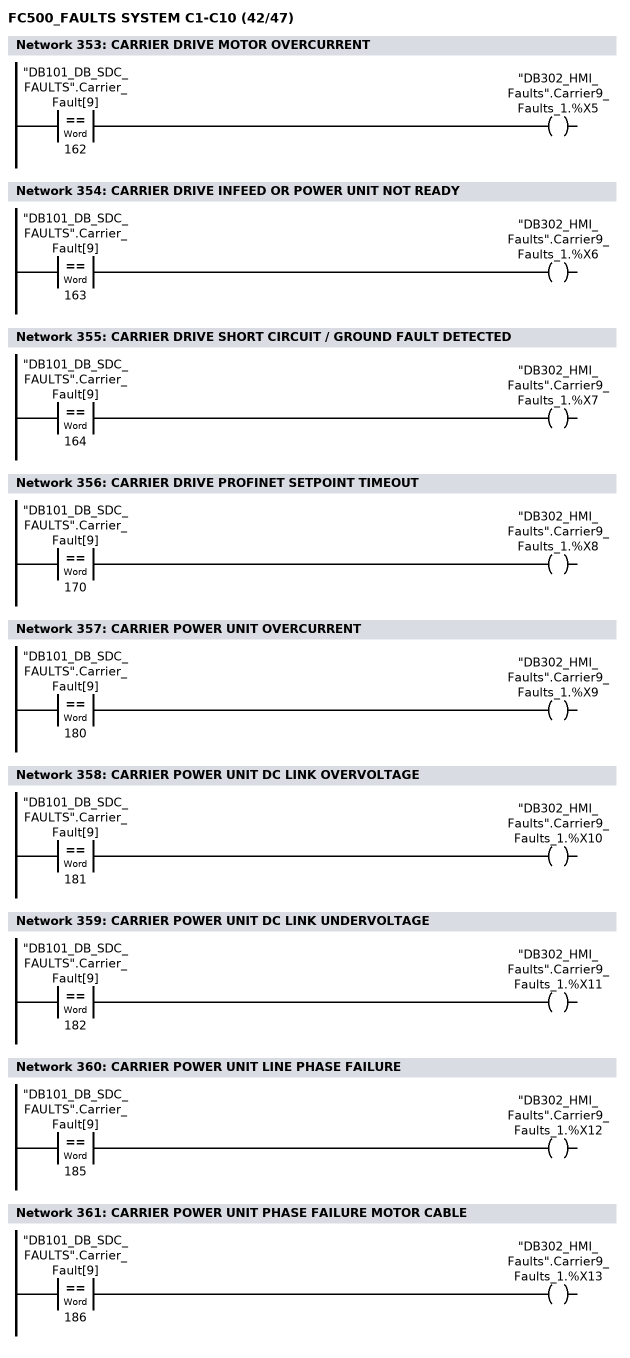
   RUNG wire#powerrail
      { S7_Templates := "SrcType := Word" } EQ_Contact(in1 := "DB101_DB_SDC_FAULTS".Carrier_Fault[9], in2 := 162)
      Coil( "DB302_HMI_Faults".Carrier9_Faults_1.%X5 )
   END_RUNG
   // the same network as SCL:
   "DB302_HMI_Faults".Carrier9_Faults_1.%X5 := "DB101_DB_SDC_FAULTS".Carrier_Fault[9] = 162;
END_REGION

REGION Network 354: CARRIER DRIVE INFEED OR POWER UNIT NOT READY
   RUNG wire#powerrail
      { S7_Templates := "SrcType := Word" } EQ_Contact(in1 := "DB101_DB_SDC_FAULTS".Carrier_Fault[9], in2 := 163)
      Coil( "DB302_HMI_Faults".Carrier9_Faults_1.%X6 )
   END_RUNG
   // the same network as SCL:
   "DB302_HMI_Faults".Carrier9_Faults_1.%X6 := "DB101_DB_SDC_FAULTS".Carrier_Fault[9] = 163;
END_REGION

REGION Network 355: CARRIER DRIVE SHORT CIRCUIT / GROUND FAULT DETECTED
   RUNG wire#powerrail
      { S7_Templates := "SrcType := Word" } EQ_Contact(in1 := "DB101_DB_SDC_FAULTS".Carrier_Fault[9], in2 := 164)
      Coil( "DB302_HMI_Faults".Carrier9_Faults_1.%X7 )
   END_RUNG
   // the same network as SCL:
   "DB302_HMI_Faults".Carrier9_Faults_1.%X7 := "DB101_DB_SDC_FAULTS".Carrier_Fault[9] = 164;
END_REGION

REGION Network 356: CARRIER DRIVE PROFINET SETPOINT TIMEOUT
   RUNG wire#powerrail
      { S7_Templates := "SrcType := Word" } EQ_Contact(in1 := "DB101_DB_SDC_FAULTS".Carrier_Fault[9], in2 := 170)
      Coil( "DB302_HMI_Faults".Carrier9_Faults_1.%X8 )
   END_RUNG
   // the same network as SCL:
   "DB302_HMI_Faults".Carrier9_Faults_1.%X8 := "DB101_DB_SDC_FAULTS".Carrier_Fault[9] = 170;
END_REGION

REGION Network 357: CARRIER POWER UNIT OVERCURRENT
   RUNG wire#powerrail
      { S7_Templates := "SrcType := Word" } EQ_Contact(in1 := "DB101_DB_SDC_FAULTS".Carrier_Fault[9], in2 := 180)
      Coil( "DB302_HMI_Faults".Carrier9_Faults_1.%X9 )
   END_RUNG
   // the same network as SCL:
   "DB302_HMI_Faults".Carrier9_Faults_1.%X9 := "DB101_DB_SDC_FAULTS".Carrier_Fault[9] = 180;
END_REGION

REGION Network 358: CARRIER POWER UNIT DC LINK OVERVOLTAGE
   RUNG wire#powerrail
      { S7_Templates := "SrcType := Word" } EQ_Contact(in1 := "DB101_DB_SDC_FAULTS".Carrier_Fault[9], in2 := 181)
      Coil( "DB302_HMI_Faults".Carrier9_Faults_1.%X10 )
   END_RUNG
   // the same network as SCL:
   "DB302_HMI_Faults".Carrier9_Faults_1.%X10 := "DB101_DB_SDC_FAULTS".Carrier_Fault[9] = 181;
END_REGION

REGION Network 359: CARRIER POWER UNIT DC LINK UNDERVOLTAGE
   RUNG wire#powerrail
      { S7_Templates := "SrcType := Word" } EQ_Contact(in1 := "DB101_DB_SDC_FAULTS".Carrier_Fault[9], in2 := 182)
      Coil( "DB302_HMI_Faults".Carrier9_Faults_1.%X11 )
   END_RUNG
   // the same network as SCL:
   "DB302_HMI_Faults".Carrier9_Faults_1.%X11 := "DB101_DB_SDC_FAULTS".Carrier_Fault[9] = 182;
END_REGION

REGION Network 360: CARRIER POWER UNIT LINE PHASE FAILURE
   RUNG wire#powerrail
      { S7_Templates := "SrcType := Word" } EQ_Contact(in1 := "DB101_DB_SDC_FAULTS".Carrier_Fault[9], in2 := 185)
      Coil( "DB302_HMI_Faults".Carrier9_Faults_1.%X12 )
   END_RUNG
   // the same network as SCL:
   "DB302_HMI_Faults".Carrier9_Faults_1.%X12 := "DB101_DB_SDC_FAULTS".Carrier_Fault[9] = 185;
END_REGION

REGION Network 361: CARRIER POWER UNIT PHASE FAILURE MOTOR CABLE
   RUNG wire#powerrail
      { S7_Templates := "SrcType := Word" } EQ_Contact(in1 := "DB101_DB_SDC_FAULTS".Carrier_Fault[9], in2 := 186)
      Coil( "DB302_HMI_Faults".Carrier9_Faults_1.%X13 )
   END_RUNG
   // the same network as SCL:
   "DB302_HMI_Faults".Carrier9_Faults_1.%X13 := "DB101_DB_SDC_FAULTS".Carrier_Fault[9] = 186;
END_REGION

REGION Network 362: CARRIER POWER UNIT GROUND FAULT
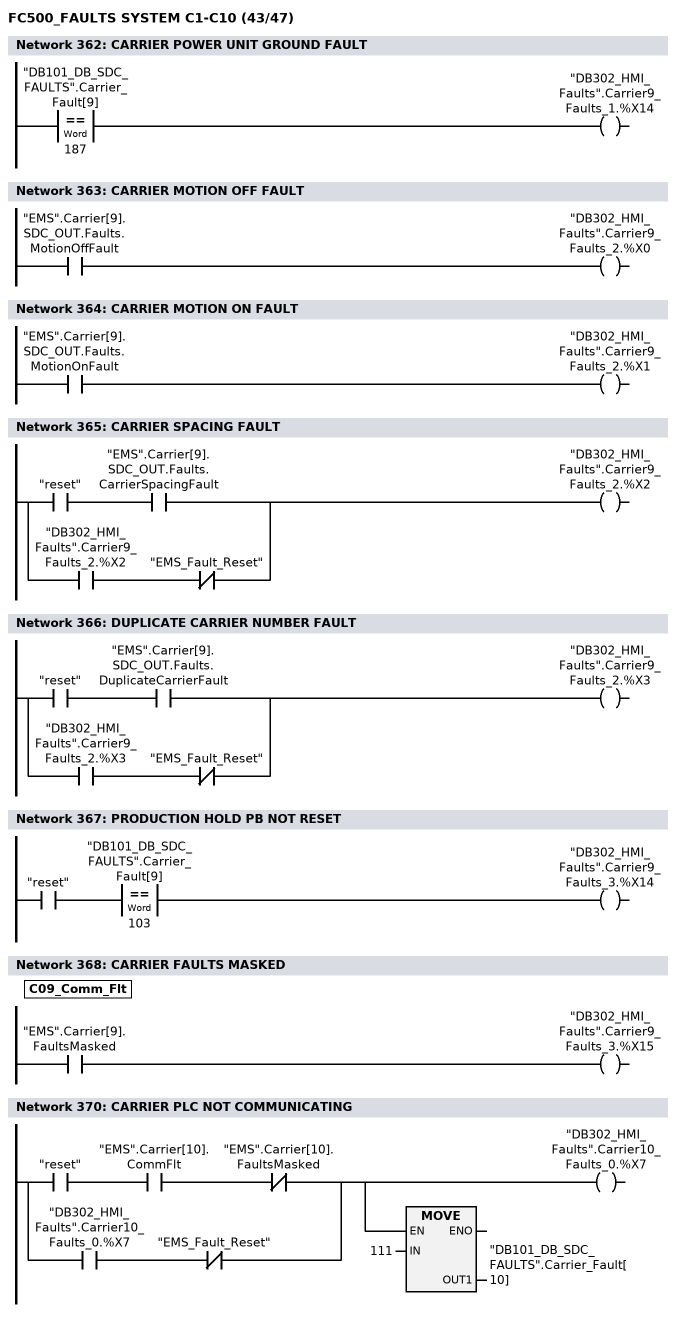
   RUNG wire#powerrail
      { S7_Templates := "SrcType := Word" } EQ_Contact(in1 := "DB101_DB_SDC_FAULTS".Carrier_Fault[9], in2 := 187)
      Coil( "DB302_HMI_Faults".Carrier9_Faults_1.%X14 )
   END_RUNG
   // the same network as SCL:
   "DB302_HMI_Faults".Carrier9_Faults_1.%X14 := "DB101_DB_SDC_FAULTS".Carrier_Fault[9] = 187;
END_REGION

REGION Network 363: CARRIER MOTION OFF FAULT
   RUNG wire#powerrail
      Contact( "EMS".Carrier[9].SDC_OUT.Faults.MotionOffFault )
      Coil( "DB302_HMI_Faults".Carrier9_Faults_2.%X0 )
   END_RUNG
   // the same network as SCL:
   "DB302_HMI_Faults".Carrier9_Faults_2.%X0 := "EMS".Carrier[9].SDC_OUT.Faults.MotionOffFault;
END_REGION

REGION Network 364: CARRIER MOTION ON FAULT
   RUNG wire#powerrail
      Contact( "EMS".Carrier[9].SDC_OUT.Faults.MotionOnFault )
      Coil( "DB302_HMI_Faults".Carrier9_Faults_2.%X1 )
   END_RUNG
   // the same network as SCL:
   "DB302_HMI_Faults".Carrier9_Faults_2.%X1 := "EMS".Carrier[9].SDC_OUT.Faults.MotionOnFault;
END_REGION

REGION Network 365: CARRIER SPACING FAULT
   RUNG wire#powerrail
      Contact( "reset" )
      Contact( "EMS".Carrier[9].SDC_OUT.Faults.CarrierSpacingFault )
      wire#w1
      Coil( "DB302_HMI_Faults".Carrier9_Faults_2.%X2 )
   END_RUNG
   RUNG wire#powerrail
      Contact( "DB302_HMI_Faults".Carrier9_Faults_2.%X2 )
      I_Contact( "EMS_Fault_Reset" )
   END_RUNG wire#w1
   // the same network as SCL:
   "DB302_HMI_Faults".Carrier9_Faults_2.%X2 := ("reset" AND "EMS".Carrier[9].SDC_OUT.Faults.CarrierSpacingFault) OR ("DB302_HMI_Faults".Carrier9_Faults_2.%X2 AND NOT "EMS_Fault_Reset");
END_REGION

REGION Network 366: DUPLICATE CARRIER NUMBER FAULT
   RUNG wire#powerrail
      Contact( "reset" )
      Contact( "EMS".Carrier[9].SDC_OUT.Faults.DuplicateCarrierFault )
      wire#w1
      Coil( "DB302_HMI_Faults".Carrier9_Faults_2.%X3 )
   END_RUNG
   RUNG wire#powerrail
      Contact( "DB302_HMI_Faults".Carrier9_Faults_2.%X3 )
      I_Contact( "EMS_Fault_Reset" )
   END_RUNG wire#w1
   // the same network as SCL:
   "DB302_HMI_Faults".Carrier9_Faults_2.%X3 := ("reset" AND "EMS".Carrier[9].SDC_OUT.Faults.DuplicateCarrierFault) OR ("DB302_HMI_Faults".Carrier9_Faults_2.%X3 AND NOT "EMS_Fault_Reset");
END_REGION

REGION Network 367: PRODUCTION HOLD PB NOT RESET
   RUNG wire#powerrail
      Contact( "reset" )
      { S7_Templates := "SrcType := Word" } EQ_Contact(in1 := "DB101_DB_SDC_FAULTS".Carrier_Fault[9], in2 := 103)
      Coil( "DB302_HMI_Faults".Carrier9_Faults_3.%X14 )
   END_RUNG
   // the same network as SCL:
   "DB302_HMI_Faults".Carrier9_Faults_3.%X14 := "reset" AND ("DB101_DB_SDC_FAULTS".Carrier_Fault[9] = 103);
END_REGION

REGION Network 368: CARRIER FAULTS MASKED
   Label( C09_Comm_Flt )
   RUNG wire#powerrail
      Contact( "EMS".Carrier[9].FaultsMasked )
      Coil( "DB302_HMI_Faults".Carrier9_Faults_3.%X15 )
   END_RUNG
   // the same network as SCL:
   C09_Comm_Flt:
   "DB302_HMI_Faults".Carrier9_Faults_3.%X15 := "EMS".Carrier[9].FaultsMasked;
END_REGION

REGION Network 369: CARRIER 10 FAULTS
END_REGION

REGION Network 370: CARRIER PLC NOT COMMUNICATING
   RUNG wire#powerrail
      Contact( "reset" )
      Contact( "EMS".Carrier[10].CommFlt )
      I_Contact( "EMS".Carrier[10].FaultsMasked )
      wire#w1
      Coil( "DB302_HMI_Faults".Carrier10_Faults_0.%X7 )
   END_RUNG
   RUNG wire#powerrail
      Contact( "DB302_HMI_Faults".Carrier10_Faults_0.%X7 )
      I_Contact( "EMS_Fault_Reset" )
   END_RUNG wire#w1
   RUNG wire#w1
      Move(in := 111, out1 => "DB101_DB_SDC_FAULTS".Carrier_Fault[10])
   END_RUNG
   // the same network as SCL:
   "DB302_HMI_Faults".Carrier10_Faults_0.%X7 := ("reset" AND "EMS".Carrier[10].CommFlt AND NOT "EMS".Carrier[10].FaultsMasked) OR ("DB302_HMI_Faults".Carrier10_Faults_0.%X7 AND NOT "EMS_Fault_Reset");
   IF "DB302_HMI_Faults".Carrier10_Faults_0.%X7 THEN "DB101_DB_SDC_FAULTS".Carrier_Fault[10] := 111; END_IF;
END_REGION

REGION Network 371
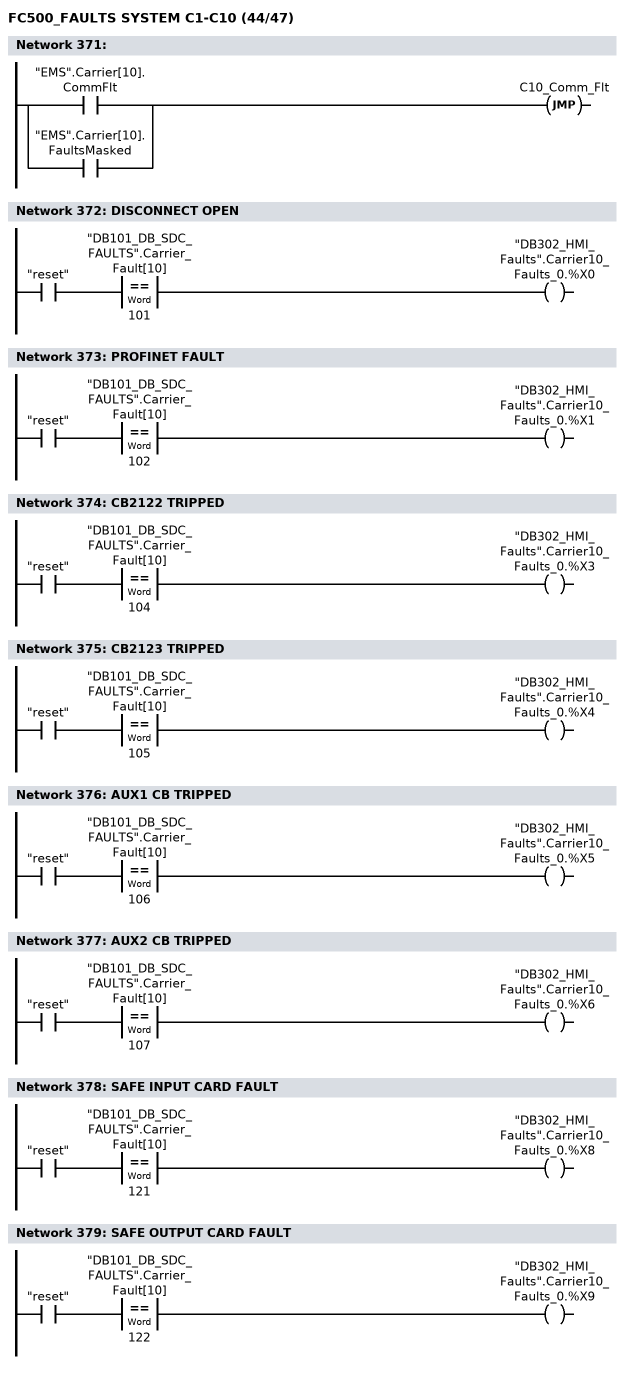
   RUNG wire#powerrail
      Contact( "EMS".Carrier[10].CommFlt )
      wire#w1
      JumpCoil( C10_Comm_Flt )
   END_RUNG
   RUNG wire#powerrail
      Contact( "EMS".Carrier[10].FaultsMasked )
   END_RUNG wire#w1
   // the same network as SCL:
   IF "EMS".Carrier[10].CommFlt OR "EMS".Carrier[10].FaultsMasked THEN GOTO C10_Comm_Flt; END_IF;
END_REGION

REGION Network 372: DISCONNECT OPEN
   RUNG wire#powerrail
      Contact( "reset" )
      { S7_Templates := "SrcType := Word" } EQ_Contact(in1 := "DB101_DB_SDC_FAULTS".Carrier_Fault[10], in2 := 101)
      Coil( "DB302_HMI_Faults".Carrier10_Faults_0.%X0 )
   END_RUNG
   // the same network as SCL:
   "DB302_HMI_Faults".Carrier10_Faults_0.%X0 := "reset" AND ("DB101_DB_SDC_FAULTS".Carrier_Fault[10] = 101);
END_REGION

REGION Network 373: PROFINET FAULT
   RUNG wire#powerrail
      Contact( "reset" )
      { S7_Templates := "SrcType := Word" } EQ_Contact(in1 := "DB101_DB_SDC_FAULTS".Carrier_Fault[10], in2 := 102)
      Coil( "DB302_HMI_Faults".Carrier10_Faults_0.%X1 )
   END_RUNG
   // the same network as SCL:
   "DB302_HMI_Faults".Carrier10_Faults_0.%X1 := "reset" AND ("DB101_DB_SDC_FAULTS".Carrier_Fault[10] = 102);
END_REGION

REGION Network 374: CB2122 TRIPPED
   RUNG wire#powerrail
      Contact( "reset" )
      { S7_Templates := "SrcType := Word" } EQ_Contact(in1 := "DB101_DB_SDC_FAULTS".Carrier_Fault[10], in2 := 104)
      Coil( "DB302_HMI_Faults".Carrier10_Faults_0.%X3 )
   END_RUNG
   // the same network as SCL:
   "DB302_HMI_Faults".Carrier10_Faults_0.%X3 := "reset" AND ("DB101_DB_SDC_FAULTS".Carrier_Fault[10] = 104);
END_REGION

REGION Network 375: CB2123 TRIPPED
   RUNG wire#powerrail
      Contact( "reset" )
      { S7_Templates := "SrcType := Word" } EQ_Contact(in1 := "DB101_DB_SDC_FAULTS".Carrier_Fault[10], in2 := 105)
      Coil( "DB302_HMI_Faults".Carrier10_Faults_0.%X4 )
   END_RUNG
   // the same network as SCL:
   "DB302_HMI_Faults".Carrier10_Faults_0.%X4 := "reset" AND ("DB101_DB_SDC_FAULTS".Carrier_Fault[10] = 105);
END_REGION

REGION Network 376: AUX1 CB TRIPPED
   RUNG wire#powerrail
      Contact( "reset" )
      { S7_Templates := "SrcType := Word" } EQ_Contact(in1 := "DB101_DB_SDC_FAULTS".Carrier_Fault[10], in2 := 106)
      Coil( "DB302_HMI_Faults".Carrier10_Faults_0.%X5 )
   END_RUNG
   // the same network as SCL:
   "DB302_HMI_Faults".Carrier10_Faults_0.%X5 := "reset" AND ("DB101_DB_SDC_FAULTS".Carrier_Fault[10] = 106);
END_REGION

REGION Network 377: AUX2 CB TRIPPED
   RUNG wire#powerrail
      Contact( "reset" )
      { S7_Templates := "SrcType := Word" } EQ_Contact(in1 := "DB101_DB_SDC_FAULTS".Carrier_Fault[10], in2 := 107)
      Coil( "DB302_HMI_Faults".Carrier10_Faults_0.%X6 )
   END_RUNG
   // the same network as SCL:
   "DB302_HMI_Faults".Carrier10_Faults_0.%X6 := "reset" AND ("DB101_DB_SDC_FAULTS".Carrier_Fault[10] = 107);
END_REGION

REGION Network 378: SAFE INPUT CARD FAULT
   RUNG wire#powerrail
      Contact( "reset" )
      { S7_Templates := "SrcType := Word" } EQ_Contact(in1 := "DB101_DB_SDC_FAULTS".Carrier_Fault[10], in2 := 121)
      Coil( "DB302_HMI_Faults".Carrier10_Faults_0.%X8 )
   END_RUNG
   // the same network as SCL:
   "DB302_HMI_Faults".Carrier10_Faults_0.%X8 := "reset" AND ("DB101_DB_SDC_FAULTS".Carrier_Fault[10] = 121);
END_REGION

REGION Network 379: SAFE OUTPUT CARD FAULT
   RUNG wire#powerrail
      Contact( "reset" )
      { S7_Templates := "SrcType := Word" } EQ_Contact(in1 := "DB101_DB_SDC_FAULTS".Carrier_Fault[10], in2 := 122)
      Coil( "DB302_HMI_Faults".Carrier10_Faults_0.%X9 )
   END_RUNG
   // the same network as SCL:
   "DB302_HMI_Faults".Carrier10_Faults_0.%X9 := "reset" AND ("DB101_DB_SDC_FAULTS".Carrier_Fault[10] = 122);
END_REGION

REGION Network 380: STANDARD INPUT CARD FAULT
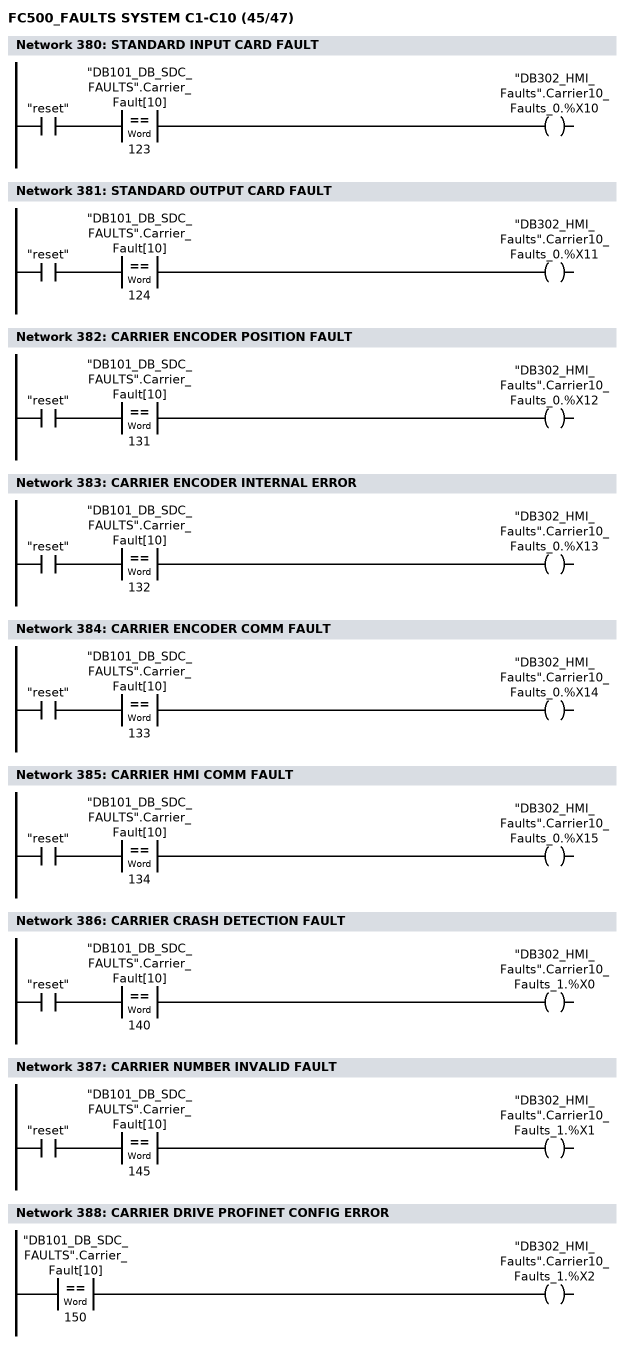
   RUNG wire#powerrail
      Contact( "reset" )
      { S7_Templates := "SrcType := Word" } EQ_Contact(in1 := "DB101_DB_SDC_FAULTS".Carrier_Fault[10], in2 := 123)
      Coil( "DB302_HMI_Faults".Carrier10_Faults_0.%X10 )
   END_RUNG
   // the same network as SCL:
   "DB302_HMI_Faults".Carrier10_Faults_0.%X10 := "reset" AND ("DB101_DB_SDC_FAULTS".Carrier_Fault[10] = 123);
END_REGION

REGION Network 381: STANDARD OUTPUT CARD FAULT
   RUNG wire#powerrail
      Contact( "reset" )
      { S7_Templates := "SrcType := Word" } EQ_Contact(in1 := "DB101_DB_SDC_FAULTS".Carrier_Fault[10], in2 := 124)
      Coil( "DB302_HMI_Faults".Carrier10_Faults_0.%X11 )
   END_RUNG
   // the same network as SCL:
   "DB302_HMI_Faults".Carrier10_Faults_0.%X11 := "reset" AND ("DB101_DB_SDC_FAULTS".Carrier_Fault[10] = 124);
END_REGION

REGION Network 382: CARRIER ENCODER POSITION FAULT
   RUNG wire#powerrail
      Contact( "reset" )
      { S7_Templates := "SrcType := Word" } EQ_Contact(in1 := "DB101_DB_SDC_FAULTS".Carrier_Fault[10], in2 := 131)
      Coil( "DB302_HMI_Faults".Carrier10_Faults_0.%X12 )
   END_RUNG
   // the same network as SCL:
   "DB302_HMI_Faults".Carrier10_Faults_0.%X12 := "reset" AND ("DB101_DB_SDC_FAULTS".Carrier_Fault[10] = 131);
END_REGION

REGION Network 383: CARRIER ENCODER INTERNAL ERROR
   RUNG wire#powerrail
      Contact( "reset" )
      { S7_Templates := "SrcType := Word" } EQ_Contact(in1 := "DB101_DB_SDC_FAULTS".Carrier_Fault[10], in2 := 132)
      Coil( "DB302_HMI_Faults".Carrier10_Faults_0.%X13 )
   END_RUNG
   // the same network as SCL:
   "DB302_HMI_Faults".Carrier10_Faults_0.%X13 := "reset" AND ("DB101_DB_SDC_FAULTS".Carrier_Fault[10] = 132);
END_REGION

REGION Network 384: CARRIER ENCODER COMM FAULT
   RUNG wire#powerrail
      Contact( "reset" )
      { S7_Templates := "SrcType := Word" } EQ_Contact(in1 := "DB101_DB_SDC_FAULTS".Carrier_Fault[10], in2 := 133)
      Coil( "DB302_HMI_Faults".Carrier10_Faults_0.%X14 )
   END_RUNG
   // the same network as SCL:
   "DB302_HMI_Faults".Carrier10_Faults_0.%X14 := "reset" AND ("DB101_DB_SDC_FAULTS".Carrier_Fault[10] = 133);
END_REGION

REGION Network 385: CARRIER HMI COMM FAULT
   RUNG wire#powerrail
      Contact( "reset" )
      { S7_Templates := "SrcType := Word" } EQ_Contact(in1 := "DB101_DB_SDC_FAULTS".Carrier_Fault[10], in2 := 134)
      Coil( "DB302_HMI_Faults".Carrier10_Faults_0.%X15 )
   END_RUNG
   // the same network as SCL:
   "DB302_HMI_Faults".Carrier10_Faults_0.%X15 := "reset" AND ("DB101_DB_SDC_FAULTS".Carrier_Fault[10] = 134);
END_REGION

REGION Network 386: CARRIER CRASH DETECTION FAULT
   RUNG wire#powerrail
      Contact( "reset" )
      { S7_Templates := "SrcType := Word" } EQ_Contact(in1 := "DB101_DB_SDC_FAULTS".Carrier_Fault[10], in2 := 140)
      Coil( "DB302_HMI_Faults".Carrier10_Faults_1.%X0 )
   END_RUNG
   // the same network as SCL:
   "DB302_HMI_Faults".Carrier10_Faults_1.%X0 := "reset" AND ("DB101_DB_SDC_FAULTS".Carrier_Fault[10] = 140);
END_REGION

REGION Network 387: CARRIER NUMBER INVALID FAULT
   RUNG wire#powerrail
      Contact( "reset" )
      { S7_Templates := "SrcType := Word" } EQ_Contact(in1 := "DB101_DB_SDC_FAULTS".Carrier_Fault[10], in2 := 145)
      Coil( "DB302_HMI_Faults".Carrier10_Faults_1.%X1 )
   END_RUNG
   // the same network as SCL:
   "DB302_HMI_Faults".Carrier10_Faults_1.%X1 := "reset" AND ("DB101_DB_SDC_FAULTS".Carrier_Fault[10] = 145);
END_REGION

REGION Network 388: CARRIER DRIVE PROFINET CONFIG ERROR
   RUNG wire#powerrail
      { S7_Templates := "SrcType := Word" } EQ_Contact(in1 := "DB101_DB_SDC_FAULTS".Carrier_Fault[10], in2 := 150)
      Coil( "DB302_HMI_Faults".Carrier10_Faults_1.%X2 )
   END_RUNG
   // the same network as SCL:
   "DB302_HMI_Faults".Carrier10_Faults_1.%X2 := "DB101_DB_SDC_FAULTS".Carrier_Fault[10] = 150;
END_REGION

REGION Network 389: CARRIER DRIVE INTERNAL COMM ERROR
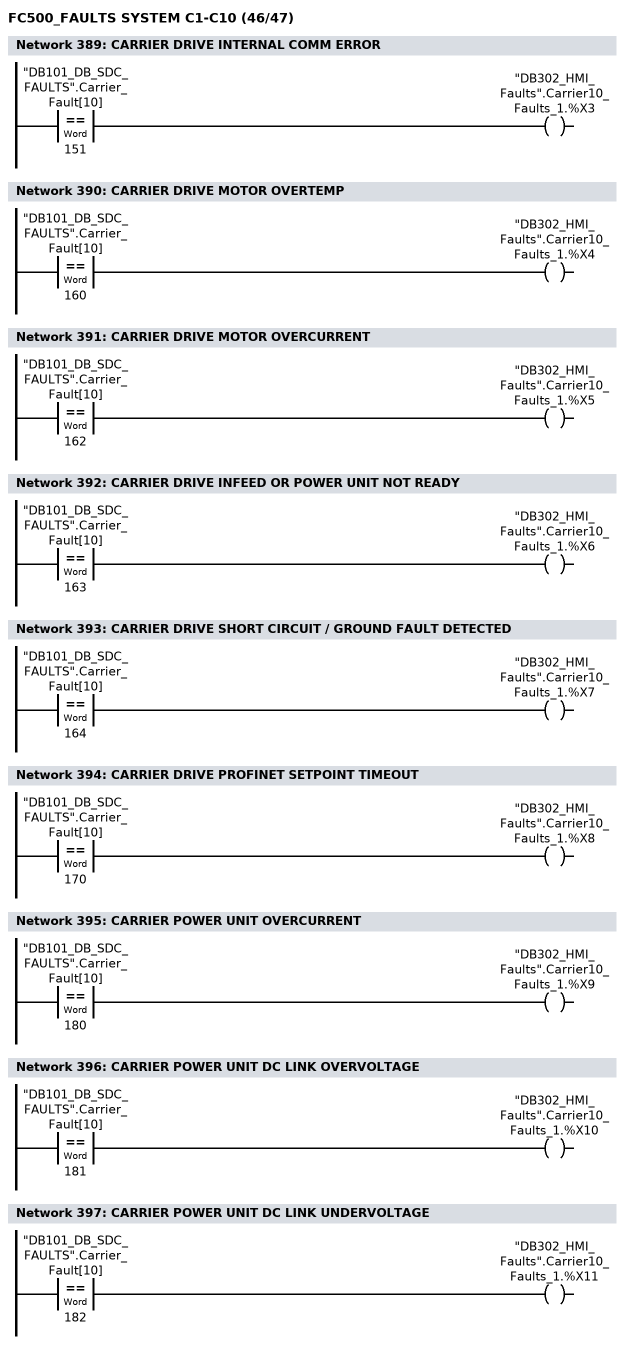
   RUNG wire#powerrail
      { S7_Templates := "SrcType := Word" } EQ_Contact(in1 := "DB101_DB_SDC_FAULTS".Carrier_Fault[10], in2 := 151)
      Coil( "DB302_HMI_Faults".Carrier10_Faults_1.%X3 )
   END_RUNG
   // the same network as SCL:
   "DB302_HMI_Faults".Carrier10_Faults_1.%X3 := "DB101_DB_SDC_FAULTS".Carrier_Fault[10] = 151;
END_REGION

REGION Network 390: CARRIER DRIVE MOTOR OVERTEMP
   RUNG wire#powerrail
      { S7_Templates := "SrcType := Word" } EQ_Contact(in1 := "DB101_DB_SDC_FAULTS".Carrier_Fault[10], in2 := 160)
      Coil( "DB302_HMI_Faults".Carrier10_Faults_1.%X4 )
   END_RUNG
   // the same network as SCL:
   "DB302_HMI_Faults".Carrier10_Faults_1.%X4 := "DB101_DB_SDC_FAULTS".Carrier_Fault[10] = 160;
END_REGION

REGION Network 391: CARRIER DRIVE MOTOR OVERCURRENT
   RUNG wire#powerrail
      { S7_Templates := "SrcType := Word" } EQ_Contact(in1 := "DB101_DB_SDC_FAULTS".Carrier_Fault[10], in2 := 162)
      Coil( "DB302_HMI_Faults".Carrier10_Faults_1.%X5 )
   END_RUNG
   // the same network as SCL:
   "DB302_HMI_Faults".Carrier10_Faults_1.%X5 := "DB101_DB_SDC_FAULTS".Carrier_Fault[10] = 162;
END_REGION

REGION Network 392: CARRIER DRIVE INFEED OR POWER UNIT NOT READY
   RUNG wire#powerrail
      { S7_Templates := "SrcType := Word" } EQ_Contact(in1 := "DB101_DB_SDC_FAULTS".Carrier_Fault[10], in2 := 163)
      Coil( "DB302_HMI_Faults".Carrier10_Faults_1.%X6 )
   END_RUNG
   // the same network as SCL:
   "DB302_HMI_Faults".Carrier10_Faults_1.%X6 := "DB101_DB_SDC_FAULTS".Carrier_Fault[10] = 163;
END_REGION

REGION Network 393: CARRIER DRIVE SHORT CIRCUIT / GROUND FAULT DETECTED
   RUNG wire#powerrail
      { S7_Templates := "SrcType := Word" } EQ_Contact(in1 := "DB101_DB_SDC_FAULTS".Carrier_Fault[10], in2 := 164)
      Coil( "DB302_HMI_Faults".Carrier10_Faults_1.%X7 )
   END_RUNG
   // the same network as SCL:
   "DB302_HMI_Faults".Carrier10_Faults_1.%X7 := "DB101_DB_SDC_FAULTS".Carrier_Fault[10] = 164;
END_REGION

REGION Network 394: CARRIER DRIVE PROFINET SETPOINT TIMEOUT
   RUNG wire#powerrail
      { S7_Templates := "SrcType := Word" } EQ_Contact(in1 := "DB101_DB_SDC_FAULTS".Carrier_Fault[10], in2 := 170)
      Coil( "DB302_HMI_Faults".Carrier10_Faults_1.%X8 )
   END_RUNG
   // the same network as SCL:
   "DB302_HMI_Faults".Carrier10_Faults_1.%X8 := "DB101_DB_SDC_FAULTS".Carrier_Fault[10] = 170;
END_REGION

REGION Network 395: CARRIER POWER UNIT OVERCURRENT
   RUNG wire#powerrail
      { S7_Templates := "SrcType := Word" } EQ_Contact(in1 := "DB101_DB_SDC_FAULTS".Carrier_Fault[10], in2 := 180)
      Coil( "DB302_HMI_Faults".Carrier10_Faults_1.%X9 )
   END_RUNG
   // the same network as SCL:
   "DB302_HMI_Faults".Carrier10_Faults_1.%X9 := "DB101_DB_SDC_FAULTS".Carrier_Fault[10] = 180;
END_REGION

REGION Network 396: CARRIER POWER UNIT DC LINK OVERVOLTAGE
   RUNG wire#powerrail
      { S7_Templates := "SrcType := Word" } EQ_Contact(in1 := "DB101_DB_SDC_FAULTS".Carrier_Fault[10], in2 := 181)
      Coil( "DB302_HMI_Faults".Carrier10_Faults_1.%X10 )
   END_RUNG
   // the same network as SCL:
   "DB302_HMI_Faults".Carrier10_Faults_1.%X10 := "DB101_DB_SDC_FAULTS".Carrier_Fault[10] = 181;
END_REGION

REGION Network 397: CARRIER POWER UNIT DC LINK UNDERVOLTAGE
   RUNG wire#powerrail
      { S7_Templates := "SrcType := Word" } EQ_Contact(in1 := "DB101_DB_SDC_FAULTS".Carrier_Fault[10], in2 := 182)
      Coil( "DB302_HMI_Faults".Carrier10_Faults_1.%X11 )
   END_RUNG
   // the same network as SCL:
   "DB302_HMI_Faults".Carrier10_Faults_1.%X11 := "DB101_DB_SDC_FAULTS".Carrier_Fault[10] = 182;
END_REGION

REGION Network 398: CARRIER POWER UNIT LINE PHASE FAILURE
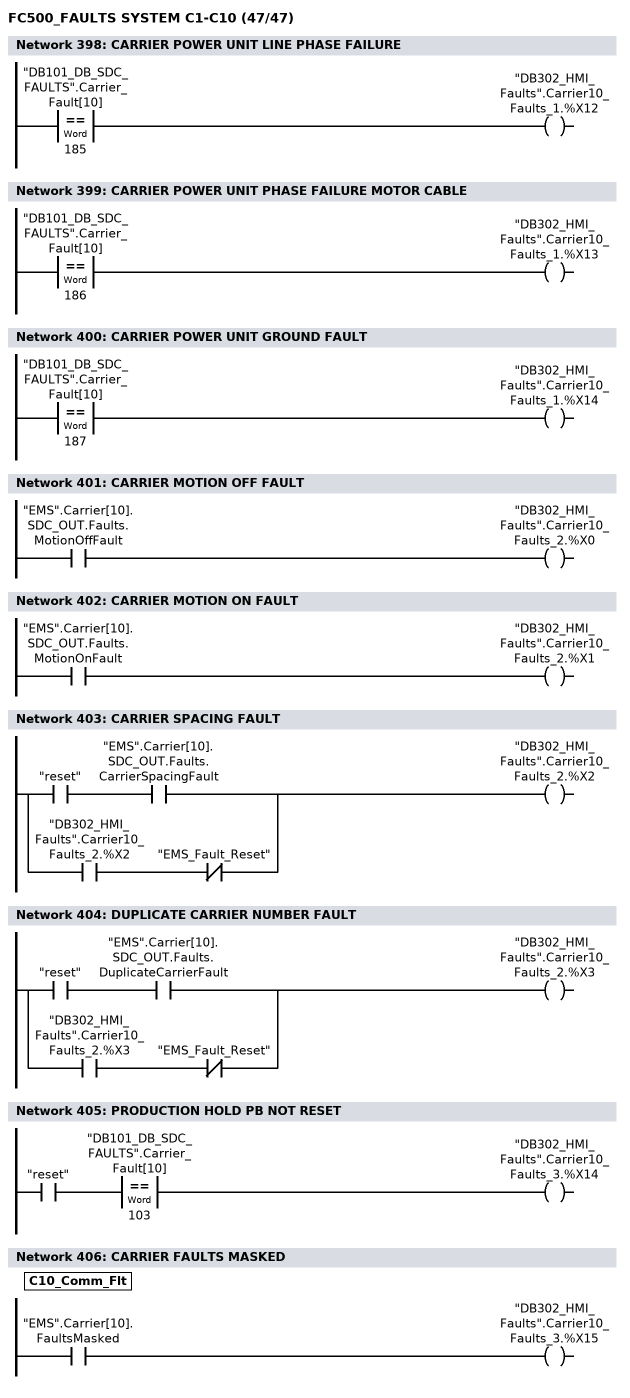
   RUNG wire#powerrail
      { S7_Templates := "SrcType := Word" } EQ_Contact(in1 := "DB101_DB_SDC_FAULTS".Carrier_Fault[10], in2 := 185)
      Coil( "DB302_HMI_Faults".Carrier10_Faults_1.%X12 )
   END_RUNG
   // the same network as SCL:
   "DB302_HMI_Faults".Carrier10_Faults_1.%X12 := "DB101_DB_SDC_FAULTS".Carrier_Fault[10] = 185;
END_REGION

REGION Network 399: CARRIER POWER UNIT PHASE FAILURE MOTOR CABLE
   RUNG wire#powerrail
      { S7_Templates := "SrcType := Word" } EQ_Contact(in1 := "DB101_DB_SDC_FAULTS".Carrier_Fault[10], in2 := 186)
      Coil( "DB302_HMI_Faults".Carrier10_Faults_1.%X13 )
   END_RUNG
   // the same network as SCL:
   "DB302_HMI_Faults".Carrier10_Faults_1.%X13 := "DB101_DB_SDC_FAULTS".Carrier_Fault[10] = 186;
END_REGION

REGION Network 400: CARRIER POWER UNIT GROUND FAULT
   RUNG wire#powerrail
      { S7_Templates := "SrcType := Word" } EQ_Contact(in1 := "DB101_DB_SDC_FAULTS".Carrier_Fault[10], in2 := 187)
      Coil( "DB302_HMI_Faults".Carrier10_Faults_1.%X14 )
   END_RUNG
   // the same network as SCL:
   "DB302_HMI_Faults".Carrier10_Faults_1.%X14 := "DB101_DB_SDC_FAULTS".Carrier_Fault[10] = 187;
END_REGION

REGION Network 401: CARRIER MOTION OFF FAULT
   RUNG wire#powerrail
      Contact( "EMS".Carrier[10].SDC_OUT.Faults.MotionOffFault )
      Coil( "DB302_HMI_Faults".Carrier10_Faults_2.%X0 )
   END_RUNG
   // the same network as SCL:
   "DB302_HMI_Faults".Carrier10_Faults_2.%X0 := "EMS".Carrier[10].SDC_OUT.Faults.MotionOffFault;
END_REGION

REGION Network 402: CARRIER MOTION ON FAULT
   RUNG wire#powerrail
      Contact( "EMS".Carrier[10].SDC_OUT.Faults.MotionOnFault )
      Coil( "DB302_HMI_Faults".Carrier10_Faults_2.%X1 )
   END_RUNG
   // the same network as SCL:
   "DB302_HMI_Faults".Carrier10_Faults_2.%X1 := "EMS".Carrier[10].SDC_OUT.Faults.MotionOnFault;
END_REGION

REGION Network 403: CARRIER SPACING FAULT
   RUNG wire#powerrail
      Contact( "reset" )
      Contact( "EMS".Carrier[10].SDC_OUT.Faults.CarrierSpacingFault )
      wire#w1
      Coil( "DB302_HMI_Faults".Carrier10_Faults_2.%X2 )
   END_RUNG
   RUNG wire#powerrail
      Contact( "DB302_HMI_Faults".Carrier10_Faults_2.%X2 )
      I_Contact( "EMS_Fault_Reset" )
   END_RUNG wire#w1
   // the same network as SCL:
   "DB302_HMI_Faults".Carrier10_Faults_2.%X2 := ("reset" AND "EMS".Carrier[10].SDC_OUT.Faults.CarrierSpacingFault) OR ("DB302_HMI_Faults".Carrier10_Faults_2.%X2 AND NOT "EMS_Fault_Reset");
END_REGION

REGION Network 404: DUPLICATE CARRIER NUMBER FAULT
   RUNG wire#powerrail
      Contact( "reset" )
      Contact( "EMS".Carrier[10].SDC_OUT.Faults.DuplicateCarrierFault )
      wire#w1
      Coil( "DB302_HMI_Faults".Carrier10_Faults_2.%X3 )
   END_RUNG
   RUNG wire#powerrail
      Contact( "DB302_HMI_Faults".Carrier10_Faults_2.%X3 )
      I_Contact( "EMS_Fault_Reset" )
   END_RUNG wire#w1
   // the same network as SCL:
   "DB302_HMI_Faults".Carrier10_Faults_2.%X3 := ("reset" AND "EMS".Carrier[10].SDC_OUT.Faults.DuplicateCarrierFault) OR ("DB302_HMI_Faults".Carrier10_Faults_2.%X3 AND NOT "EMS_Fault_Reset");
END_REGION

REGION Network 405: PRODUCTION HOLD PB NOT RESET
   RUNG wire#powerrail
      Contact( "reset" )
      { S7_Templates := "SrcType := Word" } EQ_Contact(in1 := "DB101_DB_SDC_FAULTS".Carrier_Fault[10], in2 := 103)
      Coil( "DB302_HMI_Faults".Carrier10_Faults_3.%X14 )
   END_RUNG
   // the same network as SCL:
   "DB302_HMI_Faults".Carrier10_Faults_3.%X14 := "reset" AND ("DB101_DB_SDC_FAULTS".Carrier_Fault[10] = 103);
END_REGION

REGION Network 406: CARRIER FAULTS MASKED
   Label( C10_Comm_Flt )
   RUNG wire#powerrail
      Contact( "EMS".Carrier[10].FaultsMasked )
      Coil( "DB302_HMI_Faults".Carrier10_Faults_3.%X15 )
   END_RUNG
   // the same network as SCL:
   C10_Comm_Flt:
   "DB302_HMI_Faults".Carrier10_Faults_3.%X15 := "EMS".Carrier[10].FaultsMasked;
END_REGION
END_FUNCTION

FUNCTION "FC501_FAULTS C11-C20" : Void   // FC501, LAD
{ S7_Optimized_Access := 'TRUE' }
VERSION : 0.1
BEGIN

REGION Network 1: CARRIER 11 FAULTS
END_REGION

REGION Network 2: CARRIER PLC NOT COMMUNICATING
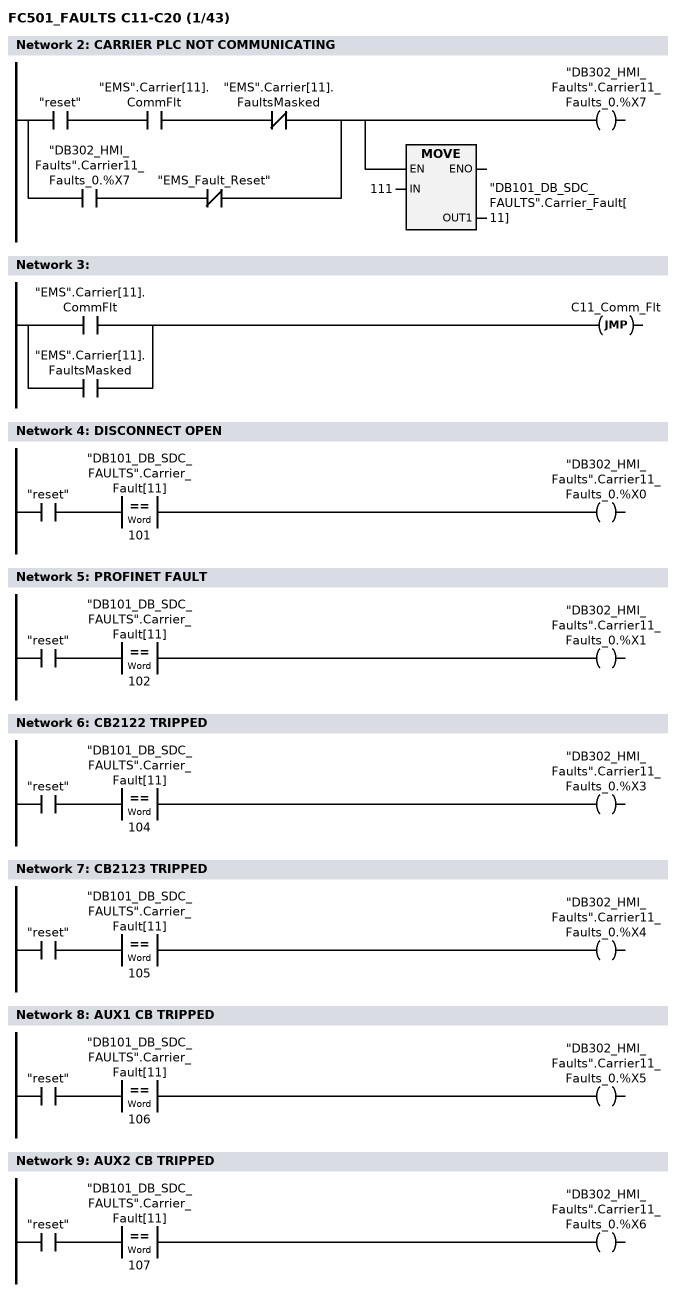
   RUNG wire#powerrail
      Contact( "reset" )
      Contact( "EMS".Carrier[11].CommFlt )
      I_Contact( "EMS".Carrier[11].FaultsMasked )
      wire#w1
      Coil( "DB302_HMI_Faults".Carrier11_Faults_0.%X7 )
   END_RUNG
   RUNG wire#powerrail
      Contact( "DB302_HMI_Faults".Carrier11_Faults_0.%X7 )
      I_Contact( "EMS_Fault_Reset" )
   END_RUNG wire#w1
   RUNG wire#w1
      Move(in := 111, out1 => "DB101_DB_SDC_FAULTS".Carrier_Fault[11])
   END_RUNG
   // the same network as SCL:
   "DB302_HMI_Faults".Carrier11_Faults_0.%X7 := ("reset" AND "EMS".Carrier[11].CommFlt AND NOT "EMS".Carrier[11].FaultsMasked) OR ("DB302_HMI_Faults".Carrier11_Faults_0.%X7 AND NOT "EMS_Fault_Reset");
   IF "DB302_HMI_Faults".Carrier11_Faults_0.%X7 THEN "DB101_DB_SDC_FAULTS".Carrier_Fault[11] := 111; END_IF;
END_REGION

REGION Network 3
   RUNG wire#powerrail
      Contact( "EMS".Carrier[11].CommFlt )
      wire#w1
      JumpCoil( C11_Comm_Flt )
   END_RUNG
   RUNG wire#powerrail
      Contact( "EMS".Carrier[11].FaultsMasked )
   END_RUNG wire#w1
   // the same network as SCL:
   IF "EMS".Carrier[11].CommFlt OR "EMS".Carrier[11].FaultsMasked THEN GOTO C11_Comm_Flt; END_IF;
END_REGION

REGION Network 4: DISCONNECT OPEN
   RUNG wire#powerrail
      Contact( "reset" )
      { S7_Templates := "SrcType := Word" } EQ_Contact(in1 := "DB101_DB_SDC_FAULTS".Carrier_Fault[11], in2 := 101)
      Coil( "DB302_HMI_Faults".Carrier11_Faults_0.%X0 )
   END_RUNG
   // the same network as SCL:
   "DB302_HMI_Faults".Carrier11_Faults_0.%X0 := "reset" AND ("DB101_DB_SDC_FAULTS".Carrier_Fault[11] = 101);
END_REGION

REGION Network 5: PROFINET FAULT
   RUNG wire#powerrail
      Contact( "reset" )
      { S7_Templates := "SrcType := Word" } EQ_Contact(in1 := "DB101_DB_SDC_FAULTS".Carrier_Fault[11], in2 := 102)
      Coil( "DB302_HMI_Faults".Carrier11_Faults_0.%X1 )
   END_RUNG
   // the same network as SCL:
   "DB302_HMI_Faults".Carrier11_Faults_0.%X1 := "reset" AND ("DB101_DB_SDC_FAULTS".Carrier_Fault[11] = 102);
END_REGION

REGION Network 6: CB2122 TRIPPED
   RUNG wire#powerrail
      Contact( "reset" )
      { S7_Templates := "SrcType := Word" } EQ_Contact(in1 := "DB101_DB_SDC_FAULTS".Carrier_Fault[11], in2 := 104)
      Coil( "DB302_HMI_Faults".Carrier11_Faults_0.%X3 )
   END_RUNG
   // the same network as SCL:
   "DB302_HMI_Faults".Carrier11_Faults_0.%X3 := "reset" AND ("DB101_DB_SDC_FAULTS".Carrier_Fault[11] = 104);
END_REGION

REGION Network 7: CB2123 TRIPPED
   RUNG wire#powerrail
      Contact( "reset" )
      { S7_Templates := "SrcType := Word" } EQ_Contact(in1 := "DB101_DB_SDC_FAULTS".Carrier_Fault[11], in2 := 105)
      Coil( "DB302_HMI_Faults".Carrier11_Faults_0.%X4 )
   END_RUNG
   // the same network as SCL:
   "DB302_HMI_Faults".Carrier11_Faults_0.%X4 := "reset" AND ("DB101_DB_SDC_FAULTS".Carrier_Fault[11] = 105);
END_REGION

REGION Network 8: AUX1 CB TRIPPED
   RUNG wire#powerrail
      Contact( "reset" )
      { S7_Templates := "SrcType := Word" } EQ_Contact(in1 := "DB101_DB_SDC_FAULTS".Carrier_Fault[11], in2 := 106)
      Coil( "DB302_HMI_Faults".Carrier11_Faults_0.%X5 )
   END_RUNG
   // the same network as SCL:
   "DB302_HMI_Faults".Carrier11_Faults_0.%X5 := "reset" AND ("DB101_DB_SDC_FAULTS".Carrier_Fault[11] = 106);
END_REGION

REGION Network 9: AUX2 CB TRIPPED
   RUNG wire#powerrail
      Contact( "reset" )
      { S7_Templates := "SrcType := Word" } EQ_Contact(in1 := "DB101_DB_SDC_FAULTS".Carrier_Fault[11], in2 := 107)
      Coil( "DB302_HMI_Faults".Carrier11_Faults_0.%X6 )
   END_RUNG
   // the same network as SCL:
   "DB302_HMI_Faults".Carrier11_Faults_0.%X6 := "reset" AND ("DB101_DB_SDC_FAULTS".Carrier_Fault[11] = 107);
END_REGION

REGION Network 10: SAFE INPUT CARD FAULT
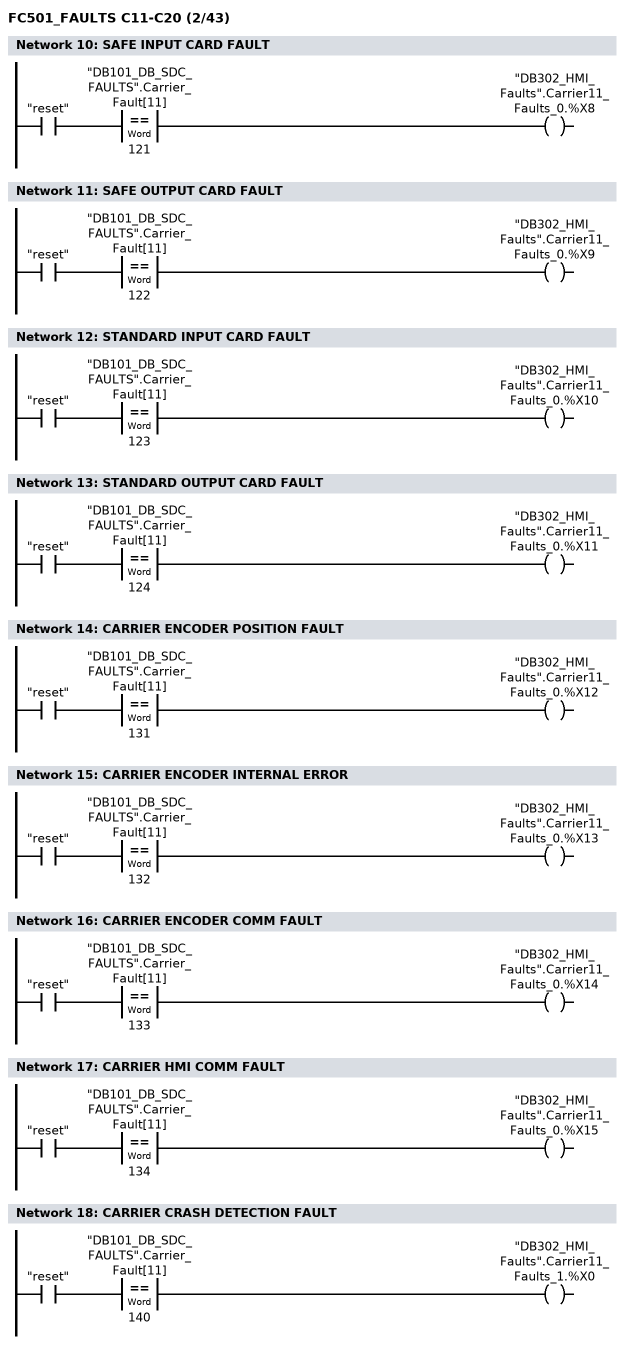
   RUNG wire#powerrail
      Contact( "reset" )
      { S7_Templates := "SrcType := Word" } EQ_Contact(in1 := "DB101_DB_SDC_FAULTS".Carrier_Fault[11], in2 := 121)
      Coil( "DB302_HMI_Faults".Carrier11_Faults_0.%X8 )
   END_RUNG
   // the same network as SCL:
   "DB302_HMI_Faults".Carrier11_Faults_0.%X8 := "reset" AND ("DB101_DB_SDC_FAULTS".Carrier_Fault[11] = 121);
END_REGION

REGION Network 11: SAFE OUTPUT CARD FAULT
   RUNG wire#powerrail
      Contact( "reset" )
      { S7_Templates := "SrcType := Word" } EQ_Contact(in1 := "DB101_DB_SDC_FAULTS".Carrier_Fault[11], in2 := 122)
      Coil( "DB302_HMI_Faults".Carrier11_Faults_0.%X9 )
   END_RUNG
   // the same network as SCL:
   "DB302_HMI_Faults".Carrier11_Faults_0.%X9 := "reset" AND ("DB101_DB_SDC_FAULTS".Carrier_Fault[11] = 122);
END_REGION

REGION Network 12: STANDARD INPUT CARD FAULT
   RUNG wire#powerrail
      Contact( "reset" )
      { S7_Templates := "SrcType := Word" } EQ_Contact(in1 := "DB101_DB_SDC_FAULTS".Carrier_Fault[11], in2 := 123)
      Coil( "DB302_HMI_Faults".Carrier11_Faults_0.%X10 )
   END_RUNG
   // the same network as SCL:
   "DB302_HMI_Faults".Carrier11_Faults_0.%X10 := "reset" AND ("DB101_DB_SDC_FAULTS".Carrier_Fault[11] = 123);
END_REGION

REGION Network 13: STANDARD OUTPUT CARD FAULT
   RUNG wire#powerrail
      Contact( "reset" )
      { S7_Templates := "SrcType := Word" } EQ_Contact(in1 := "DB101_DB_SDC_FAULTS".Carrier_Fault[11], in2 := 124)
      Coil( "DB302_HMI_Faults".Carrier11_Faults_0.%X11 )
   END_RUNG
   // the same network as SCL:
   "DB302_HMI_Faults".Carrier11_Faults_0.%X11 := "reset" AND ("DB101_DB_SDC_FAULTS".Carrier_Fault[11] = 124);
END_REGION

REGION Network 14: CARRIER ENCODER POSITION FAULT
   RUNG wire#powerrail
      Contact( "reset" )
      { S7_Templates := "SrcType := Word" } EQ_Contact(in1 := "DB101_DB_SDC_FAULTS".Carrier_Fault[11], in2 := 131)
      Coil( "DB302_HMI_Faults".Carrier11_Faults_0.%X12 )
   END_RUNG
   // the same network as SCL:
   "DB302_HMI_Faults".Carrier11_Faults_0.%X12 := "reset" AND ("DB101_DB_SDC_FAULTS".Carrier_Fault[11] = 131);
END_REGION

REGION Network 15: CARRIER ENCODER INTERNAL ERROR
   RUNG wire#powerrail
      Contact( "reset" )
      { S7_Templates := "SrcType := Word" } EQ_Contact(in1 := "DB101_DB_SDC_FAULTS".Carrier_Fault[11], in2 := 132)
      Coil( "DB302_HMI_Faults".Carrier11_Faults_0.%X13 )
   END_RUNG
   // the same network as SCL:
   "DB302_HMI_Faults".Carrier11_Faults_0.%X13 := "reset" AND ("DB101_DB_SDC_FAULTS".Carrier_Fault[11] = 132);
END_REGION

REGION Network 16: CARRIER ENCODER COMM FAULT
   RUNG wire#powerrail
      Contact( "reset" )
      { S7_Templates := "SrcType := Word" } EQ_Contact(in1 := "DB101_DB_SDC_FAULTS".Carrier_Fault[11], in2 := 133)
      Coil( "DB302_HMI_Faults".Carrier11_Faults_0.%X14 )
   END_RUNG
   // the same network as SCL:
   "DB302_HMI_Faults".Carrier11_Faults_0.%X14 := "reset" AND ("DB101_DB_SDC_FAULTS".Carrier_Fault[11] = 133);
END_REGION

REGION Network 17: CARRIER HMI COMM FAULT
   RUNG wire#powerrail
      Contact( "reset" )
      { S7_Templates := "SrcType := Word" } EQ_Contact(in1 := "DB101_DB_SDC_FAULTS".Carrier_Fault[11], in2 := 134)
      Coil( "DB302_HMI_Faults".Carrier11_Faults_0.%X15 )
   END_RUNG
   // the same network as SCL:
   "DB302_HMI_Faults".Carrier11_Faults_0.%X15 := "reset" AND ("DB101_DB_SDC_FAULTS".Carrier_Fault[11] = 134);
END_REGION
